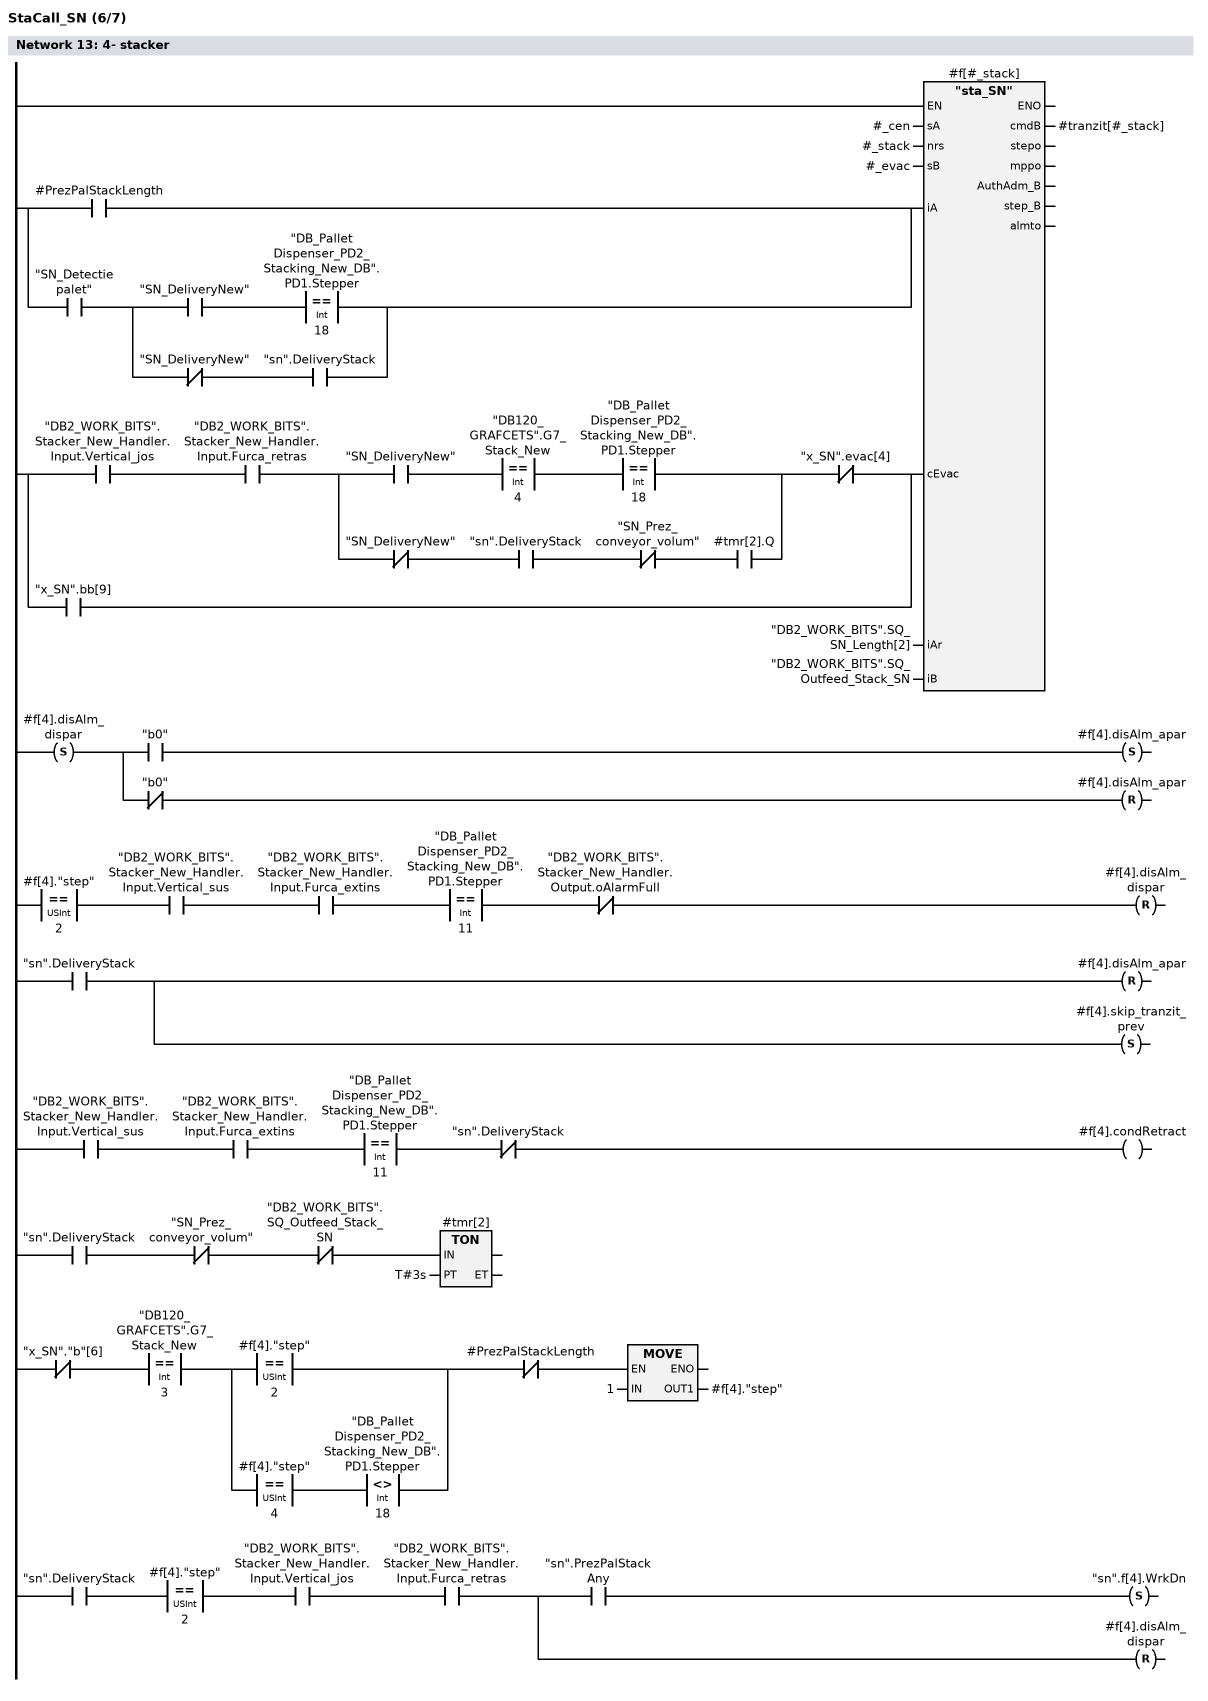
   #f[#_stack](sA := #_cen,   // "sta_SN"
               nrs := #_stack,
               sB := #_evac,
               iA := #PrezPalStackLength OR ("SN_Detectie palet" AND (("SN_DeliveryNew" AND ("DB_PalletDispenser_PD2_Stacking_New_DB".PD1.Stepper = 18)) OR (NOT "SN_DeliveryNew" AND "sn".DeliveryStack))),
               cEvac := ("DB2_WORK_BITS".Stacker_New_Handler.Input.Vertical_jos AND "DB2_WORK_BITS".Stacker_New_Handler.Input.Furca_retras AND (("SN_DeliveryNew" AND ("DB120_GRAFCETS".G7_Stack_New = 4) AND ("DB_PalletDispenser_PD2_Stacking_New_DB".PD1.Stepper = 18)) OR (NOT "SN_DeliveryNew" AND "sn".DeliveryStack AND NOT "SN_Prez_conveyor_volum" AND #tmr[2].Q)) AND NOT "x_SN".evac[4]) OR "x_SN".bb[9],
               iAr := "DB2_WORK_BITS".SQ_SN_Length[2],
               iB := "DB2_WORK_BITS".SQ_Outfeed_Stack_SN,
               cmdB => #tranzit[#_stack]);
   #f[4].disAlm_dispar := TRUE;
   IF "b0" THEN #f[4].disAlm_apar := TRUE; END_IF;
   IF NOT "b0" THEN #f[4].disAlm_apar := FALSE; END_IF;
   IF (#f[4]."step" = 2) AND "DB2_WORK_BITS".Stacker_New_Handler.Input.Vertical_sus AND "DB2_WORK_BITS".Stacker_New_Handler.Input.Furca_extins AND ("DB_PalletDispenser_PD2_Stacking_New_DB".PD1.Stepper = 11) AND NOT "DB2_WORK_BITS".Stacker_New_Handler.Output.oAlarmFull THEN
       #f[4].disAlm_dispar := FALSE;
   END_IF;
   IF "sn".DeliveryStack THEN
       #f[4].disAlm_apar := FALSE;
       #f[4].skip_tranzit_prev := TRUE;
   END_IF;
   #f[4].condRetract := "DB2_WORK_BITS".Stacker_New_Handler.Input.Vertical_sus AND "DB2_WORK_BITS".Stacker_New_Handler.Input.Furca_extins AND ("DB_PalletDispenser_PD2_Stacking_New_DB".PD1.Stepper = 11) AND NOT "sn".DeliveryStack;
   #tmr[2].TON(IN := "sn".DeliveryStack AND NOT "SN_Prez_conveyor_volum" AND NOT "DB2_WORK_BITS".SQ_Outfeed_Stack_SN,
               PT := T#3s);
   IF NOT "x_SN"."b"[6] AND ("DB120_GRAFCETS".G7_Stack_New = 3) AND ((#f[4]."step" = 2) OR ((#f[4]."step" = 4) AND ("DB_PalletDispenser_PD2_Stacking_New_DB".PD1.Stepper <> 18))) AND NOT #PrezPalStackLength THEN
       #f[4]."step" := 1;
   END_IF;
   #_w1 := "sn".DeliveryStack AND (#f[4]."step" = 2) AND "DB2_WORK_BITS".Stacker_New_Handler.Input.Vertical_jos AND "DB2_WORK_BITS".Stacker_New_Handler.Input.Furca_retras;
   IF #_w1 AND "sn".PrezPalStackAny THEN "sn".f[4].WrkDn := TRUE; END_IF;
   IF #_w1 THEN #f[4].disAlm_dispar := FALSE; END_IF;
END_REGION

REGION Network 14: 5- evac
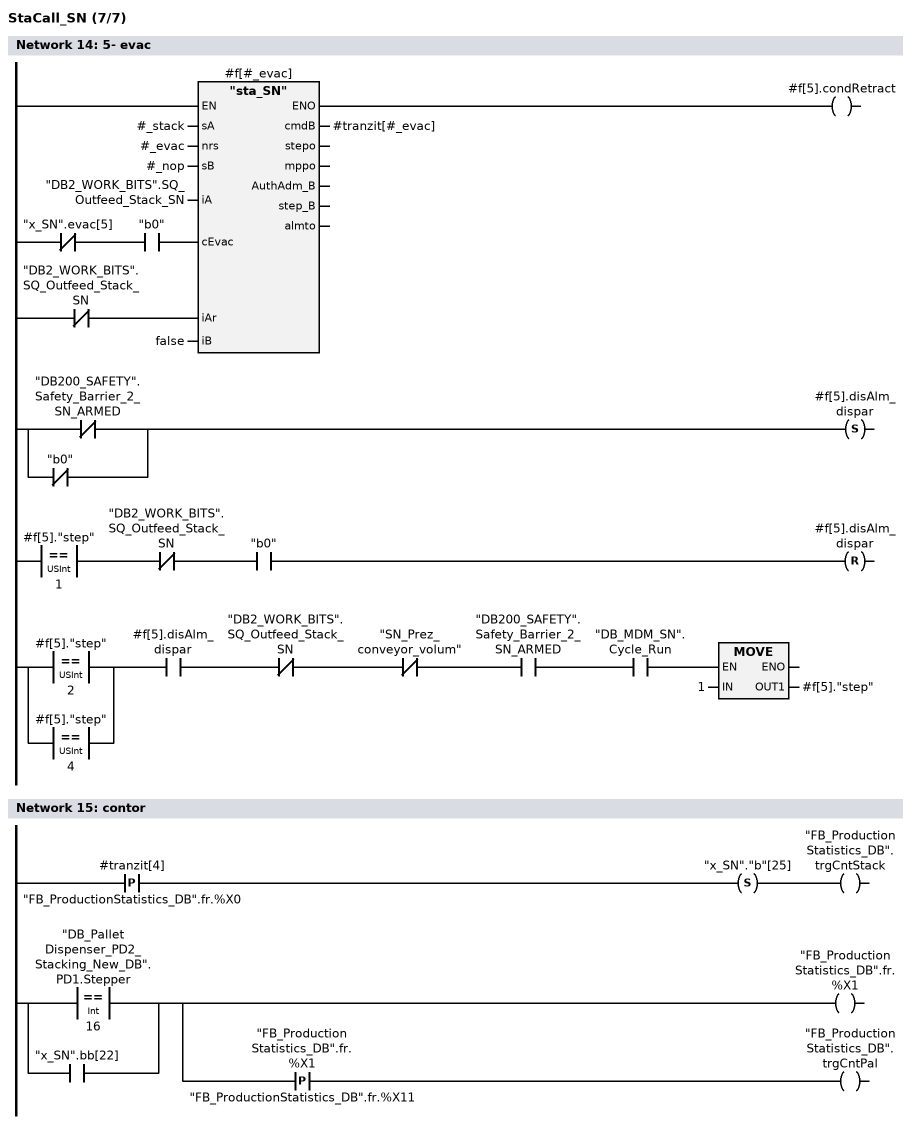
   RUNG wire#powerrail
      #f[#_evac](cEvac := wire#w1, iAr := wire#w2, sA := #_stack, nrs := #_evac, sB := #_nop, iA := "DB2_WORK_BITS".SQ_Outfeed_Stack_SN, iB := false, cmdB => #tranzit[#_evac], stepo =>, mppo =>, AuthAdm_B =>, step_B =>, almto =>)
      Coil( #f[5].condRetract )
   END_RUNG
   RUNG wire#powerrail
      I_Contact( "x_SN".evac[5] )
      Contact( "b0" )
   END_RUNG wire#w1
   RUNG wire#powerrail
      I_Contact( "DB2_WORK_BITS".SQ_Outfeed_Stack_SN )
   END_RUNG wire#w2
   RUNG wire#powerrail
      I_Contact( "DB200_SAFETY".Safety_Barrier_2_SN_ARMED )
      wire#w3
      S_Coil( #f[5].disAlm_dispar )
   END_RUNG
   RUNG wire#powerrail
      I_Contact( "b0" )
   END_RUNG wire#w3
   RUNG wire#powerrail
      { S7_Templates := "SrcType := USInt" } EQ_Contact(in1 := #f[5]."step", in2 := 1)
      I_Contact( "DB2_WORK_BITS".SQ_Outfeed_Stack_SN )
      Contact( "b0" )
      R_Coil( #f[5].disAlm_dispar )
   END_RUNG
   RUNG wire#powerrail
      { S7_Templates := "SrcType := USInt" } EQ_Contact(in1 := #f[5]."step", in2 := 2)
      wire#w4
      Contact( #f[5].disAlm_dispar )
      I_Contact( "DB2_WORK_BITS".SQ_Outfeed_Stack_SN )
      I_Contact( "SN_Prez_conveyor_volum" )
      Contact( "DB200_SAFETY".Safety_Barrier_2_SN_ARMED )
      Contact( "DB_MDM_SN".Cycle_Run )
      Move(in := 1, out1 => #f[5]."step")
   END_RUNG
   RUNG wire#powerrail
      { S7_Templates := "SrcType := USInt" } EQ_Contact(in1 := #f[5]."step", in2 := 4)
   END_RUNG wire#w4
   // the same network as SCL:
   #f[#_evac](sA := #_stack,   // "sta_SN"
              nrs := #_evac,
              sB := #_nop,
              iA := "DB2_WORK_BITS".SQ_Outfeed_Stack_SN,
              cEvac := NOT "x_SN".evac[5] AND "b0",
              iAr := NOT "DB2_WORK_BITS".SQ_Outfeed_Stack_SN,
              iB := false,
              cmdB => #tranzit[#_evac],
              ENO => #_w1);
   #f[5].condRetract := #_w1;
   IF NOT "DB200_SAFETY".Safety_Barrier_2_SN_ARMED OR NOT "b0" THEN #f[5].disAlm_dispar := TRUE; END_IF;
   IF (#f[5]."step" = 1) AND NOT "DB2_WORK_BITS".SQ_Outfeed_Stack_SN AND "b0" THEN
       #f[5].disAlm_dispar := FALSE;
   END_IF;
   IF ((#f[5]."step" = 2) OR (#f[5]."step" = 4)) AND #f[5].disAlm_dispar AND NOT "DB2_WORK_BITS".SQ_Outfeed_Stack_SN AND NOT "SN_Prez_conveyor_volum" AND "DB200_SAFETY".Safety_Barrier_2_SN_ARMED AND "DB_MDM_SN".Cycle_Run THEN
       #f[5]."step" := 1;
   END_IF;
END_REGION

REGION Network 15: contor
   RUNG wire#powerrail
      P_Contact(operand := #tranzit[4], bit := "FB_ProductionStatistics_DB".fr.%X0)
      S_Coil( "x_SN"."b"[25] )
      Coil( "FB_ProductionStatistics_DB".trgCntStack )
   END_RUNG
   RUNG wire#powerrail
      { S7_Templates := "SrcType := Int" } EQ_Contact(in1 := "DB_PalletDispenser_PD2_Stacking_New_DB".PD1.Stepper, in2 := 16)
      wire#w1
      Coil( "FB_ProductionStatistics_DB".fr.%X1 )
   END_RUNG
   RUNG wire#powerrail
      Contact( "x_SN".bb[22] )
   END_RUNG wire#w1
   RUNG wire#w1
      P_Contact(operand := "FB_ProductionStatistics_DB".fr.%X1, bit := "FB_ProductionStatistics_DB".fr.%X11)
      Coil( "FB_ProductionStatistics_DB".trgCntPal )
   END_RUNG
   // the same network as SCL:
   #_w1 := #tranzit[4] AND NOT "FB_ProductionStatistics_DB".fr.%X0;   // rising edge of #tranzit[4]
   "FB_ProductionStatistics_DB".fr.%X0 := #tranzit[4];
   IF #_w1 THEN "x_SN"."b"[25] := TRUE; END_IF;
   "FB_ProductionStatistics_DB".trgCntStack := #_w1;
   "FB_ProductionStatistics_DB".fr.%X1 := ("DB_PalletDispenser_PD2_Stacking_New_DB".PD1.Stepper = 16) OR "x_SN".bb[22];
   #_w2 := "FB_ProductionStatistics_DB".fr.%X1 AND "FB_ProductionStatistics_DB".fr.%X1 AND NOT "FB_ProductionStatistics_DB".fr.%X11;   // rising edge of "FB_ProductionStatistics_DB".fr.%X1
   "FB_ProductionStatistics_DB".fr.%X11 := "FB_ProductionStatistics_DB".fr.%X1;
   "FB_ProductionStatistics_DB".trgCntPal := #_w2;
END_REGION
END_FUNCTION_BLOCK

FUNCTION_BLOCK "sta_SN"   // FB16, LAD
{ S7_Optimized_Access := 'TRUE' }
VERSION : 0.1
   VAR_INPUT
      sA : USInt;   // statie Admit
      nrs : USInt;   // statie crt
      sB : USInt;   // statie Evac
      iA : Bool;   // conditie Admit
      cEvac : Bool;
      iAr : Bool;   // cond Release
      iB : Bool;   // cond Evac
   END_VAR
   VAR_OUTPUT
      cmdB : Bool;
      stepo : USInt;
      mppo : Bool;
      AuthAdm_B : Bool;
      step_B : USInt;
      almto : USInt;
   END_VAR
   VAR
      "step" : USInt;
      stepv : USInt;
      mpp : Bool;
      alm_apar : Bool;
      alm_disapear : Bool;
      alm_tmt : Bool;
      alm_release : Bool;
      AuthAdmit : Bool;
      AuthEvacEx : Bool;
      almt : Bool;
      WrkDn : Bool;
      condRetract : Bool;
      skip_tranzit_prev : Bool;
      product_disapear_confirmed : Bool;
      transit_end_confirmed : Bool;
      tim_alm : Array[1..6] of IEC_TIMER;
      HMI_stat_s : USInt;
      disAlm_Tmt : Bool;
      disAlm_dispar : Bool;
      disAlm_apar : Bool;
      disAlmRls : Bool;
      HMI_stat_t : USInt;
      tranzit_mem : Bool;
      cycle : Bool;
      almw : Word;
      HMI_statT : USInt;
      HMI_statS : USInt;
      tr : USInt;
      AlarmW : Word;
   END_VAR
   VAR_TEMP
      tmpui : SInt;
   END_VAR
   VAR CONSTANT
      b0 : Bool;
   END_VAR
   VAR_TEMP   // added for the SCL form of the ladder/FBD networks
      _w1 : Bool;
      _w2 : Bool;
      _w3 : Bool;
   END_VAR
BEGIN

REGION Network 1: first cycle
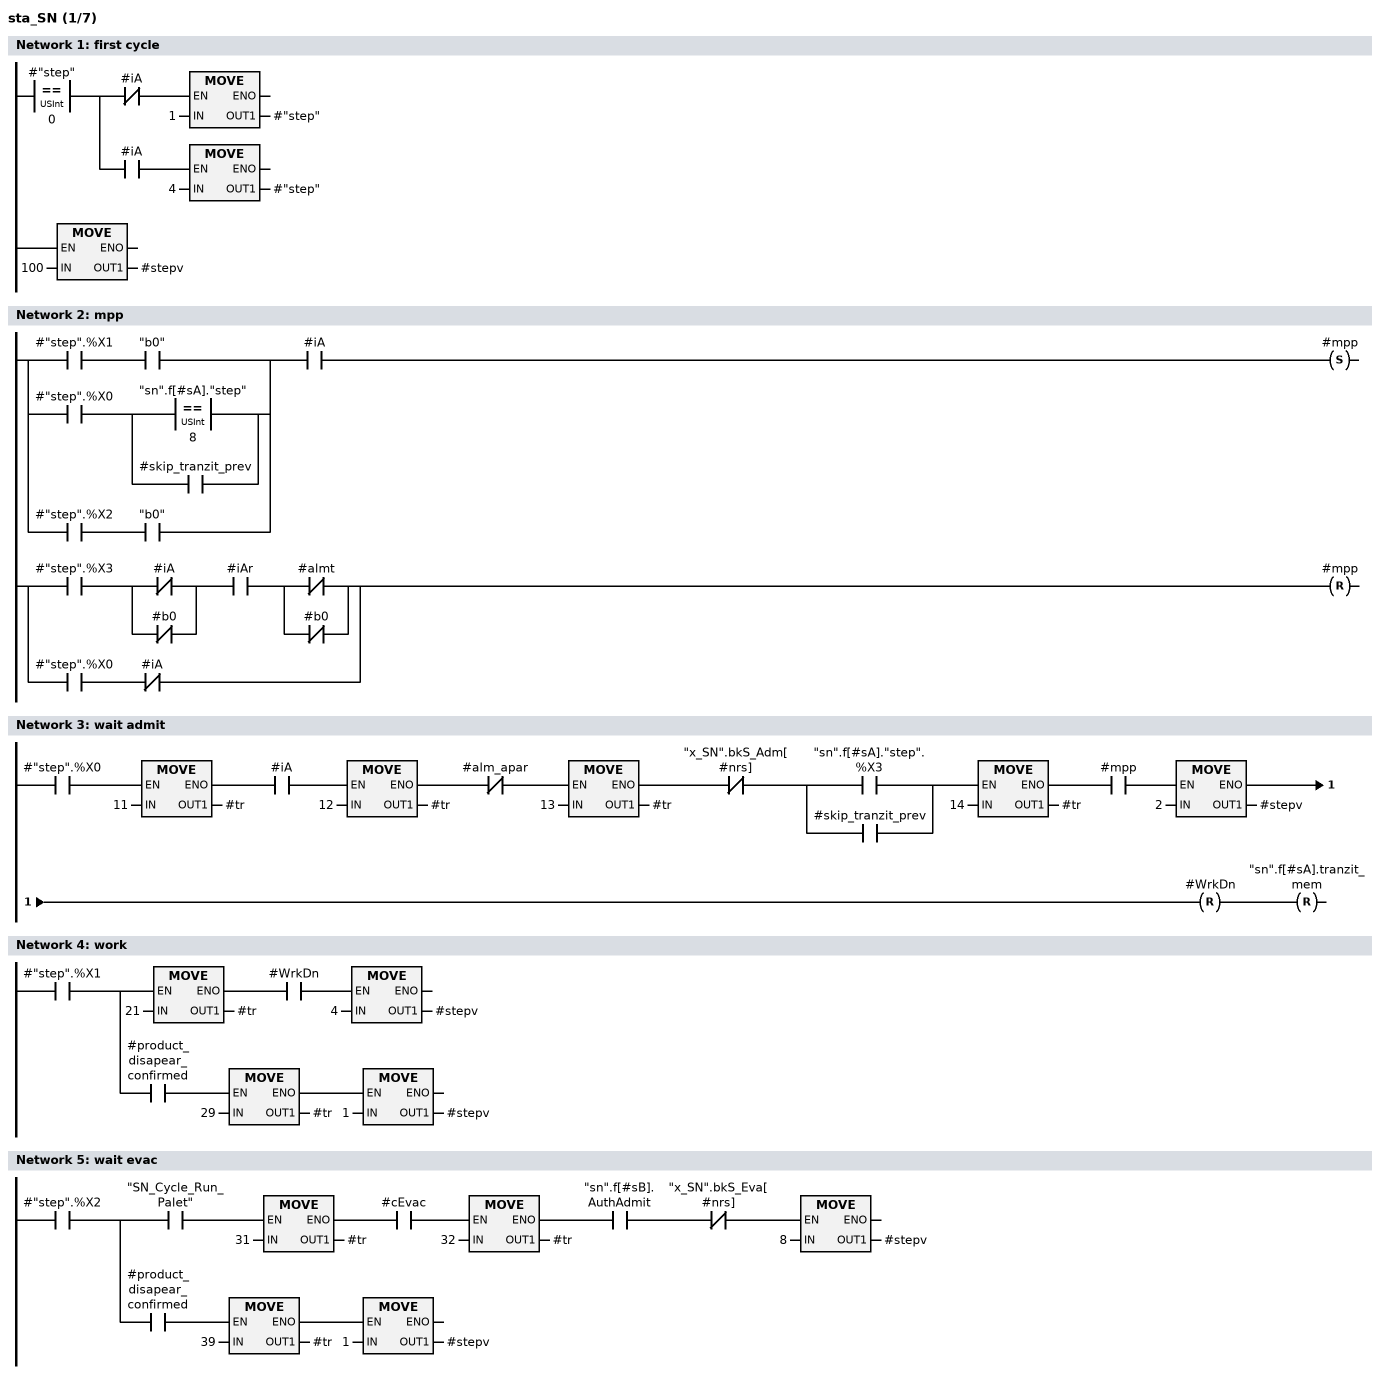
   RUNG wire#powerrail
      { S7_Templates := "SrcType := USInt" } EQ_Contact(in1 := #"step", in2 := 0)
      wire#w1
      I_Contact( #iA )
      Move(in := 1, out1 => #"step")
   END_RUNG
   RUNG wire#w1
      Contact( #iA )
      Move(in := 4, out1 => #"step")
   END_RUNG
   RUNG wire#powerrail
      Move(in := 100, out1 => #stepv)
   END_RUNG
   // the same network as SCL:
   #_w1 := #"step" = 0;
   IF #_w1 AND NOT #iA THEN #"step" := 1; END_IF;
   IF #_w1 AND #iA THEN #"step" := 4; END_IF;
   #stepv := 100;
END_REGION

REGION Network 2: mpp
   RUNG wire#powerrail
      Contact( #"step".%X1 )
      Contact( "b0" )
      wire#w1
      Contact( #iA )
      S_Coil( #mpp )
   END_RUNG
   RUNG wire#powerrail
      Contact( #"step".%X0 )
      wire#w2
      { S7_Templates := "SrcType := USInt" } EQ_Contact(in1 := "sn".f[#sA]."step", in2 := 8)
   END_RUNG wire#w1
   RUNG wire#w2
      Contact( #skip_tranzit_prev )
   END_RUNG wire#w1
   RUNG wire#powerrail
      Contact( #"step".%X2 )
      Contact( "b0" )
   END_RUNG wire#w1
   RUNG wire#powerrail
      Contact( #"step".%X3 )
      wire#w3
      I_Contact( #iA )
      wire#w4
      Contact( #iAr )
      wire#w5
      I_Contact( #almt )
      wire#w6
      R_Coil( #mpp )
   END_RUNG
   RUNG wire#w3
      I_Contact( #b0 )
   END_RUNG wire#w4
   RUNG wire#w5
      I_Contact( #b0 )
   END_RUNG wire#w6
   RUNG wire#powerrail
      Contact( #"step".%X0 )
      I_Contact( #iA )
   END_RUNG wire#w6
   // the same network as SCL:
   IF ((#"step".%X1 AND "b0") OR (#"step".%X0 AND (("sn".f[#sA]."step" = 8) OR #skip_tranzit_prev)) OR (#"step".%X2 AND "b0")) AND #iA THEN
       #mpp := TRUE;
   END_IF;
   IF (#"step".%X3 AND (NOT #iA OR NOT #b0) AND #iAr AND (NOT #almt OR NOT #b0)) OR (#"step".%X0 AND NOT #iA) THEN
       #mpp := FALSE;
   END_IF;
END_REGION

REGION Network 3: wait admit
   RUNG wire#powerrail
      Contact( #"step".%X0 )
      Move(in := 11, out1 => #tr)
      Contact( #iA )
      Move(in := 12, out1 => #tr)
      I_Contact( #alm_apar )
      Move(in := 13, out1 => #tr)
      I_Contact( "x_SN".bkS_Adm[#nrs] )
      wire#w1
      Contact( "sn".f[#sA]."step".%X3 )
      wire#w2
      Move(in := 14, out1 => #tr)
      Contact( #mpp )
      Move(in := 2, out1 => #stepv)
      R_Coil( #WrkDn )
      R_Coil( "sn".f[#sA].tranzit_mem )
   END_RUNG
   RUNG wire#w1
      Contact( #skip_tranzit_prev )
   END_RUNG wire#w2
   // the same network as SCL:
   IF #"step".%X0 THEN #tr := 11; END_IF;
   #_w1 := #"step".%X0 AND #iA;
   IF #_w1 THEN #tr := 12; END_IF;
   #_w2 := #_w1 AND NOT #alm_apar;
   IF #_w2 THEN #tr := 13; END_IF;
   #_w3 := #_w2 AND NOT "x_SN".bkS_Adm[#nrs] AND ("sn".f[#sA]."step".%X3 OR #skip_tranzit_prev);
   IF #_w3 THEN #tr := 14; END_IF;
   IF #_w3 AND #mpp THEN
       #stepv := 2;
       #WrkDn := FALSE;
       "sn".f[#sA].tranzit_mem := FALSE;
   END_IF;
END_REGION

REGION Network 4: work
   RUNG wire#powerrail
      Contact( #"step".%X1 )
      wire#w1
      Move(in := 21, out1 => #tr)
      Contact( #WrkDn )
      Move(in := 4, out1 => #stepv)
   END_RUNG
   RUNG wire#w1
      Contact( #product_disapear_confirmed )
      Move(in := 29, out1 => #tr)
      Move(in := 1, out1 => #stepv)
   END_RUNG
   // the same network as SCL:
   IF #"step".%X1 THEN #tr := 21; END_IF;
   IF #"step".%X1 AND #WrkDn THEN #stepv := 4; END_IF;
   IF #"step".%X1 AND #product_disapear_confirmed THEN
       #tr := 29;
       #stepv := 1;
   END_IF;
END_REGION

REGION Network 5: wait evac
   RUNG wire#powerrail
      Contact( #"step".%X2 )
      wire#w1
      Contact( "SN_Cycle_Run_Palet" )
      Move(in := 31, out1 => #tr)
      Contact( #cEvac )
      Move(in := 32, out1 => #tr)
      Contact( "sn".f[#sB].AuthAdmit )
      I_Contact( "x_SN".bkS_Eva[#nrs] )
      Move(in := 8, out1 => #stepv)
   END_RUNG
   RUNG wire#w1
      Contact( #product_disapear_confirmed )
      Move(in := 39, out1 => #tr)
      Move(in := 1, out1 => #stepv)
   END_RUNG
   // the same network as SCL:
   #_w1 := #"step".%X2 AND "SN_Cycle_Run_Palet";
   IF #_w1 THEN #tr := 31; END_IF;
   #_w2 := #_w1 AND #cEvac;
   IF #_w2 THEN #tr := 32; END_IF;
   IF #_w2 AND "sn".f[#sB].AuthAdmit AND NOT "x_SN".bkS_Eva[#nrs] THEN #stepv := 8; END_IF;
   IF #"step".%X2 AND #product_disapear_confirmed THEN
       #tr := 39;
       #stepv := 1;
   END_IF;
END_REGION

REGION Network 6: evac
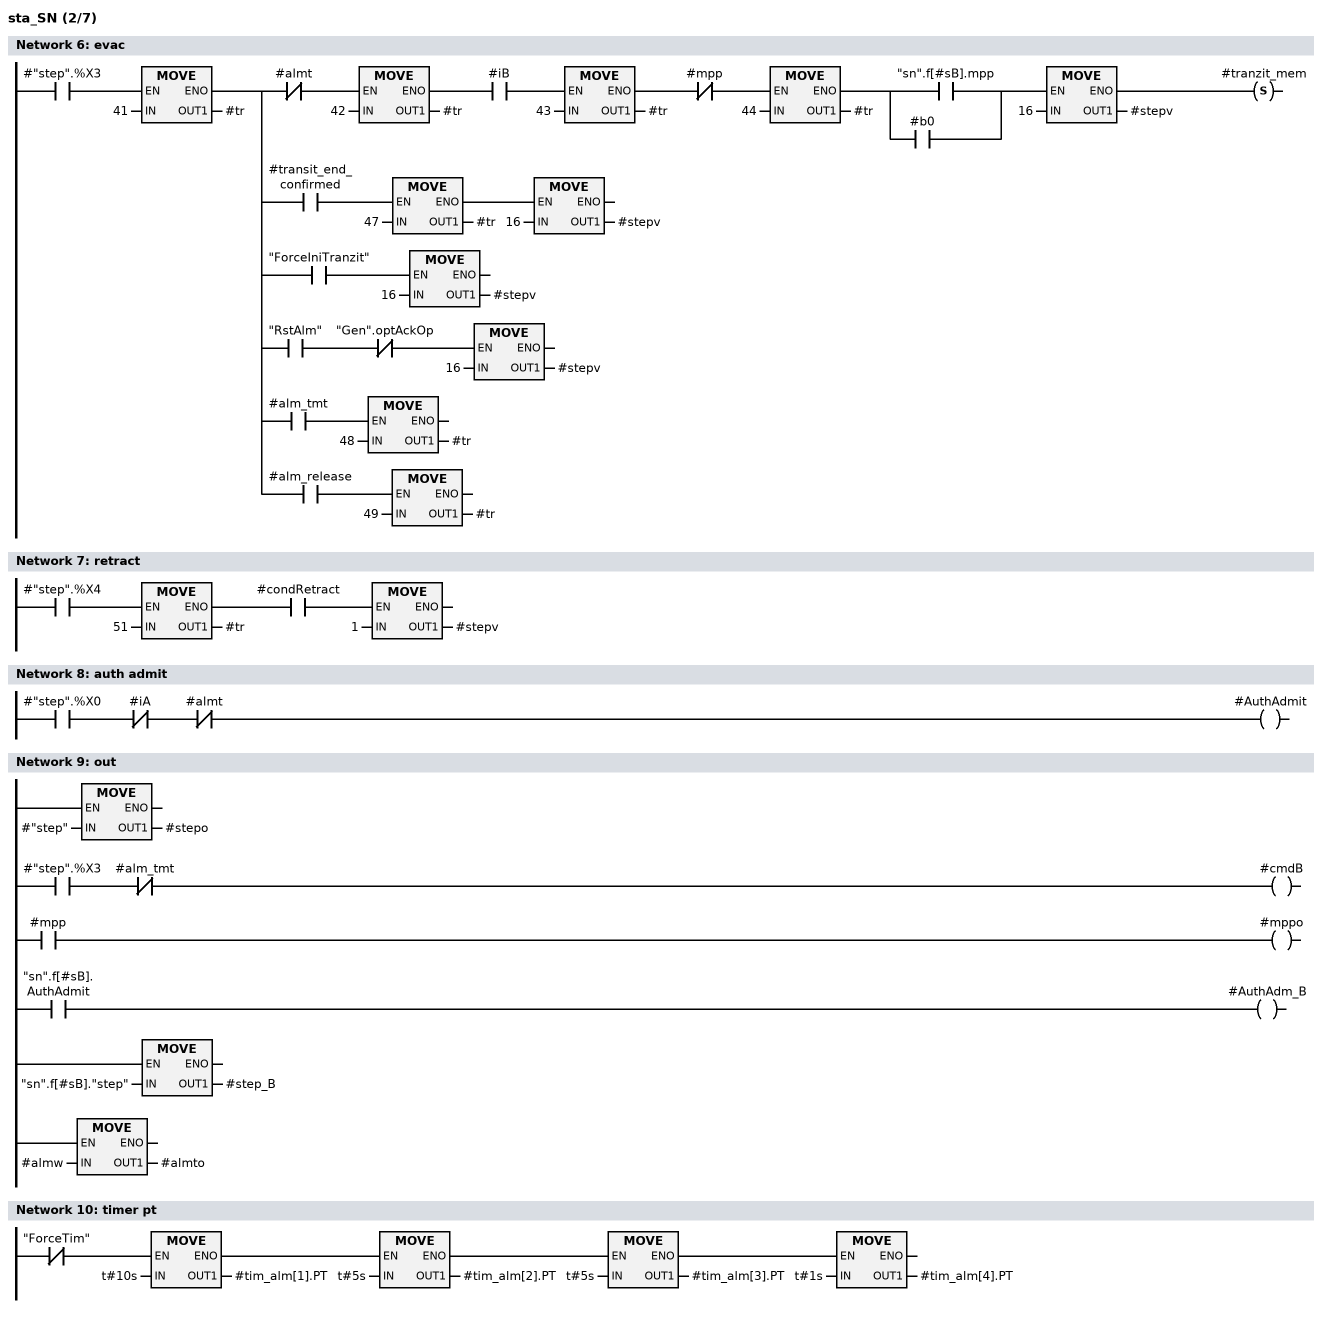
   RUNG wire#powerrail
      Contact( #"step".%X3 )
      Move(in := 41, out1 => #tr)
      wire#w1
      I_Contact( #almt )
      Move(in := 42, out1 => #tr)
      Contact( #iB )
      Move(in := 43, out1 => #tr)
      I_Contact( #mpp )
      Move(in := 44, out1 => #tr)
      wire#w2
      Contact( "sn".f[#sB].mpp )
      wire#w3
      Move(in := 16, out1 => #stepv)
      S_Coil( #tranzit_mem )
   END_RUNG
   RUNG wire#w2
      Contact( #b0 )
   END_RUNG wire#w3
   RUNG wire#w1
      Contact( #transit_end_confirmed )
      Move(in := 47, out1 => #tr)
      Move(in := 16, out1 => #stepv)
   END_RUNG
   RUNG wire#w1
      Contact( "ForceIniTranzit" )
      Move(in := 16, out1 => #stepv)
   END_RUNG
   RUNG wire#w1
      Contact( "RstAlm" )
      I_Contact( "Gen".optAckOp )
      Move(in := 16, out1 => #stepv)
   END_RUNG
   RUNG wire#w1
      Contact( #alm_tmt )
      Move(in := 48, out1 => #tr)
   END_RUNG
   RUNG wire#w1
      Contact( #alm_release )
      Move(in := 49, out1 => #tr)
   END_RUNG
   // the same network as SCL:
   IF #"step".%X3 THEN #tr := 41; END_IF;
   #_w1 := #"step".%X3 AND NOT #almt;
   IF #_w1 THEN #tr := 42; END_IF;
   #_w2 := #_w1 AND #iB;
   IF #_w2 THEN #tr := 43; END_IF;
   #_w3 := #_w2 AND NOT #mpp;
   IF #_w3 THEN #tr := 44; END_IF;
   IF #_w3 AND ("sn".f[#sB].mpp OR #b0) THEN
       #stepv := 16;
       #tranzit_mem := TRUE;
   END_IF;
   IF #"step".%X3 AND #transit_end_confirmed THEN
       #tr := 47;
       #stepv := 16;
   END_IF;
   IF #"step".%X3 AND "ForceIniTranzit" THEN #stepv := 16; END_IF;
   IF #"step".%X3 AND "RstAlm" AND NOT "Gen".optAckOp THEN #stepv := 16; END_IF;
   IF #"step".%X3 AND #alm_tmt THEN #tr := 48; END_IF;
   IF #"step".%X3 AND #alm_release THEN #tr := 49; END_IF;
END_REGION

REGION Network 7: retract
   RUNG wire#powerrail
      Contact( #"step".%X4 )
      Move(in := 51, out1 => #tr)
      Contact( #condRetract )
      Move(in := 1, out1 => #stepv)
   END_RUNG
   // the same network as SCL:
   IF #"step".%X4 THEN #tr := 51; END_IF;
   IF #"step".%X4 AND #condRetract THEN #stepv := 1; END_IF;
END_REGION

REGION Network 8: auth admit
   RUNG wire#powerrail
      Contact( #"step".%X0 )
      I_Contact( #iA )
      I_Contact( #almt )
      Coil( #AuthAdmit )
   END_RUNG
   // the same network as SCL:
   #AuthAdmit := #"step".%X0 AND NOT #iA AND NOT #almt;
END_REGION

REGION Network 9: out
   RUNG wire#powerrail
      Move(in := #"step", out1 => #stepo)
   END_RUNG
   RUNG wire#powerrail
      Contact( #"step".%X3 )
      I_Contact( #alm_tmt )
      Coil( #cmdB )
   END_RUNG
   RUNG wire#powerrail
      Contact( #mpp )
      Coil( #mppo )
   END_RUNG
   RUNG wire#powerrail
      Contact( "sn".f[#sB].AuthAdmit )
      Coil( #AuthAdm_B )
   END_RUNG
   RUNG wire#powerrail
      Move(in := "sn".f[#sB]."step", out1 => #step_B)
   END_RUNG
   RUNG wire#powerrail
      Move(in := #almw, out1 => #almto)
   END_RUNG
   // the same network as SCL:
   #stepo := #"step";
   #cmdB := #"step".%X3 AND NOT #alm_tmt;
   #mppo := #mpp;
   #AuthAdm_B := "sn".f[#sB].AuthAdmit;
   #step_B := "sn".f[#sB]."step";
   #almto := #almw;
END_REGION

REGION Network 10: timer pt
   RUNG wire#powerrail
      I_Contact( "ForceTim" )
      Move(in := t#10s, out1 => #tim_alm[1].PT)
      Move(in := t#5s, out1 => #tim_alm[2].PT)
      Move(in := t#5s, out1 => #tim_alm[3].PT)
      Move(in := t#1s, out1 => #tim_alm[4].PT)
   END_RUNG
   // the same network as SCL:
   IF NOT "ForceTim" THEN
       #tim_alm[1].PT := t#10s;
       #tim_alm[2].PT := t#5s;
       #tim_alm[3].PT := t#5s;
       #tim_alm[4].PT := t#1s;
   END_IF;
END_REGION

REGION Network 11: rst all
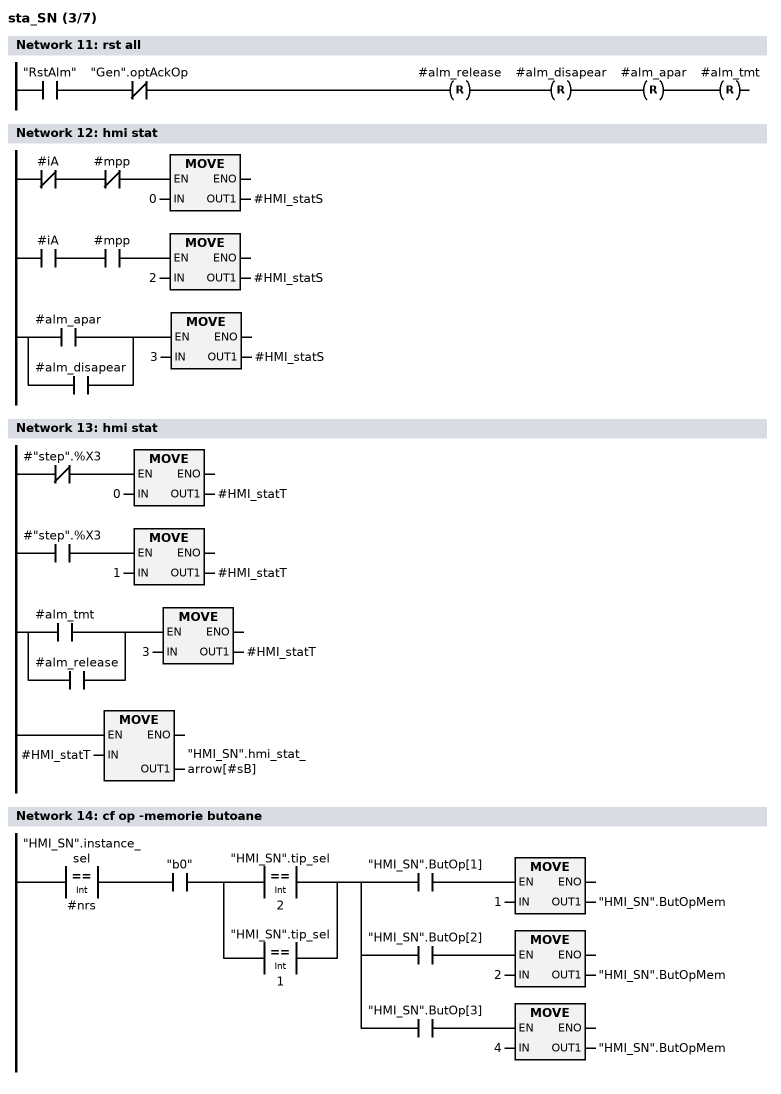
   RUNG wire#powerrail
      Contact( "RstAlm" )
      I_Contact( "Gen".optAckOp )
      R_Coil( #alm_release )
      R_Coil( #alm_disapear )
      R_Coil( #alm_apar )
      R_Coil( #alm_tmt )
   END_RUNG
   // the same network as SCL:
   IF "RstAlm" AND NOT "Gen".optAckOp THEN
       #alm_release := FALSE;
       #alm_disapear := FALSE;
       #alm_apar := FALSE;
       #alm_tmt := FALSE;
   END_IF;
END_REGION

REGION Network 12: hmi stat
   RUNG wire#powerrail
      I_Contact( #iA )
      I_Contact( #mpp )
      Move(in := 0, out1 => #HMI_statS)
   END_RUNG
   RUNG wire#powerrail
      Contact( #iA )
      Contact( #mpp )
      Move(in := 2, out1 => #HMI_statS)
   END_RUNG
   RUNG wire#powerrail
      Contact( #alm_apar )
      wire#w1
      Move(in := 3, out1 => #HMI_statS)
   END_RUNG
   RUNG wire#powerrail
      Contact( #alm_disapear )
   END_RUNG wire#w1
   // the same network as SCL:
   IF NOT #iA AND NOT #mpp THEN #HMI_statS := 0; END_IF;
   IF #iA AND #mpp THEN #HMI_statS := 2; END_IF;
   IF #alm_apar OR #alm_disapear THEN #HMI_statS := 3; END_IF;
END_REGION

REGION Network 13: hmi stat
   RUNG wire#powerrail
      I_Contact( #"step".%X3 )
      Move(in := 0, out1 => #HMI_statT)
   END_RUNG
   RUNG wire#powerrail
      Contact( #"step".%X3 )
      Move(in := 1, out1 => #HMI_statT)
   END_RUNG
   RUNG wire#powerrail
      Contact( #alm_tmt )
      wire#w1
      Move(in := 3, out1 => #HMI_statT)
   END_RUNG
   RUNG wire#powerrail
      Contact( #alm_release )
   END_RUNG wire#w1
   RUNG wire#powerrail
      Move(in := #HMI_statT, out1 => "HMI_SN".hmi_stat_arrow[#sB])
   END_RUNG
   // the same network as SCL:
   IF NOT #"step".%X3 THEN #HMI_statT := 0; END_IF;
   IF #"step".%X3 THEN #HMI_statT := 1; END_IF;
   IF #alm_tmt OR #alm_release THEN #HMI_statT := 3; END_IF;
   "HMI_SN".hmi_stat_arrow[#sB] := #HMI_statT;
END_REGION

REGION Network 14: cf op -memorie butoane
   RUNG wire#powerrail
      { S7_Templates := "SrcType := Int" } EQ_Contact(in1 := "HMI_SN".instance_sel, in2 := #nrs)
      Contact( "b0" )
      wire#w1
      { S7_Templates := "SrcType := Int" } EQ_Contact(in1 := "HMI_SN".tip_sel, in2 := 2)
      wire#w2
      Contact( "HMI_SN".ButOp[1] )
      Move(in := 1, out1 => "HMI_SN".ButOpMem)
   END_RUNG
   RUNG wire#w1
      { S7_Templates := "SrcType := Int" } EQ_Contact(in1 := "HMI_SN".tip_sel, in2 := 1)
   END_RUNG wire#w2
   RUNG wire#w2
      Contact( "HMI_SN".ButOp[2] )
      Move(in := 2, out1 => "HMI_SN".ButOpMem)
   END_RUNG
   RUNG wire#w2
      Contact( "HMI_SN".ButOp[3] )
      Move(in := 4, out1 => "HMI_SN".ButOpMem)
   END_RUNG
   // the same network as SCL:
   #_w1 := ("HMI_SN".instance_sel = #nrs) AND "b0" AND (("HMI_SN".tip_sel = 2) OR ("HMI_SN".tip_sel = 1));
   IF #_w1 AND "HMI_SN".ButOp[1] THEN "HMI_SN".ButOpMem := 1; END_IF;
   IF #_w1 AND "HMI_SN".ButOp[2] THEN "HMI_SN".ButOpMem := 2; END_IF;
   IF #_w1 AND "HMI_SN".ButOp[3] THEN "HMI_SN".ButOpMem := 4; END_IF;
END_REGION

REGION Network 15: cf op alm tmt / release
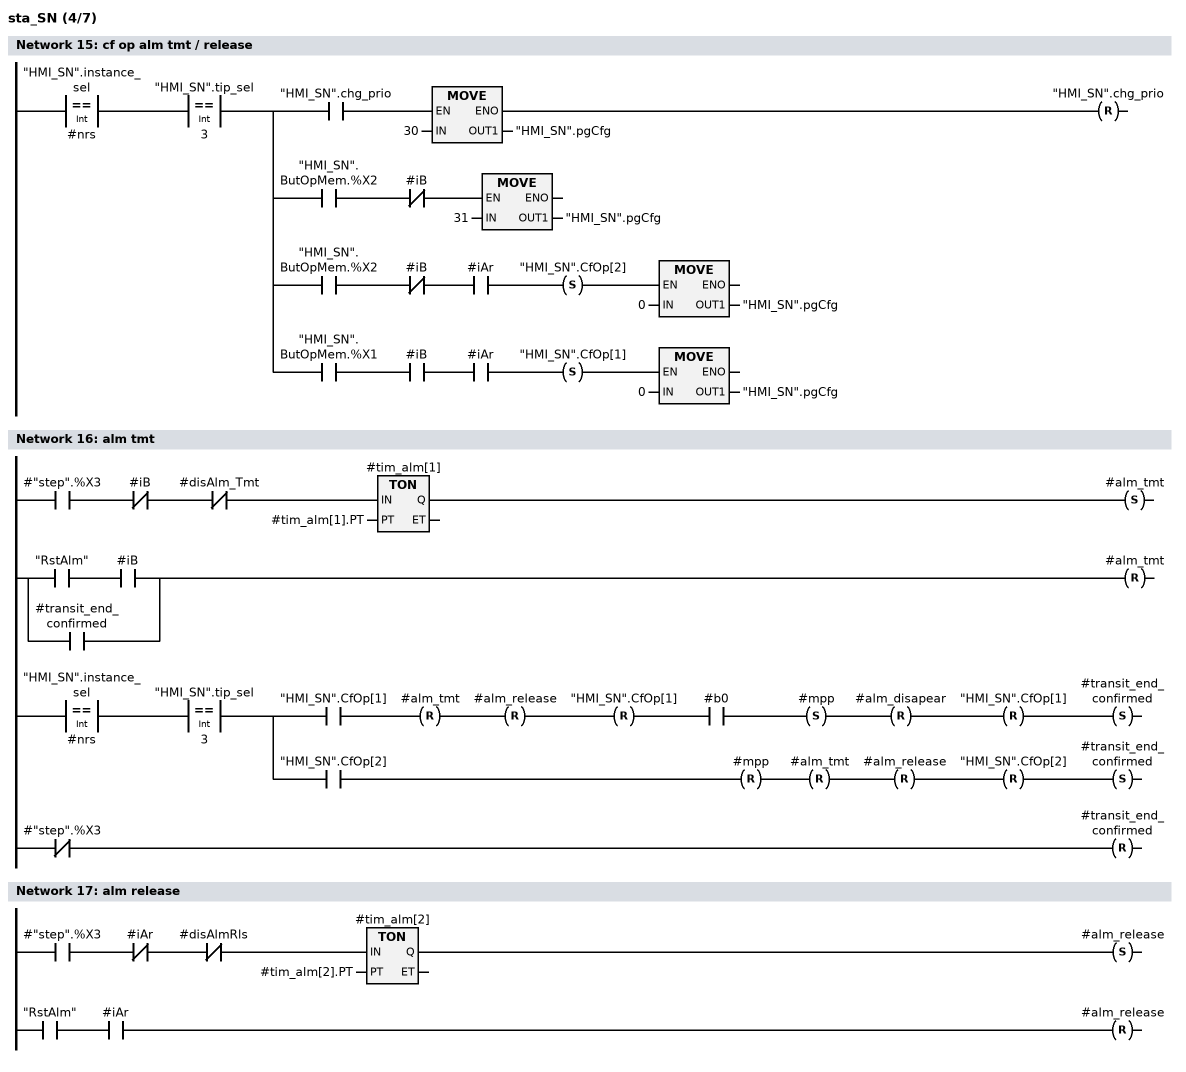
   RUNG wire#powerrail
      { S7_Templates := "SrcType := Int" } EQ_Contact(in1 := "HMI_SN".instance_sel, in2 := #nrs)
      { S7_Templates := "SrcType := Int" } EQ_Contact(in1 := "HMI_SN".tip_sel, in2 := 3)
      wire#w1
      Contact( "HMI_SN".chg_prio )
      Move(in := 30, out1 => "HMI_SN".pgCfg)
      R_Coil( "HMI_SN".chg_prio )
   END_RUNG
   RUNG wire#w1
      Contact( "HMI_SN".ButOpMem.%X2 )
      I_Contact( #iB )
      Move(in := 31, out1 => "HMI_SN".pgCfg)
   END_RUNG
   RUNG wire#w1
      Contact( "HMI_SN".ButOpMem.%X2 )
      I_Contact( #iB )
      Contact( #iAr )
      S_Coil( "HMI_SN".CfOp[2] )
      Move(in := 0, out1 => "HMI_SN".pgCfg)
   END_RUNG
   RUNG wire#w1
      Contact( "HMI_SN".ButOpMem.%X1 )
      Contact( #iB )
      Contact( #iAr )
      S_Coil( "HMI_SN".CfOp[1] )
      Move(in := 0, out1 => "HMI_SN".pgCfg)
   END_RUNG
   // the same network as SCL:
   #_w1 := ("HMI_SN".instance_sel = #nrs) AND ("HMI_SN".tip_sel = 3);
   IF #_w1 AND "HMI_SN".chg_prio THEN
       "HMI_SN".pgCfg := 30;
       "HMI_SN".chg_prio := FALSE;
   END_IF;
   IF #_w1 AND "HMI_SN".ButOpMem.%X2 AND NOT #iB THEN "HMI_SN".pgCfg := 31; END_IF;
   IF #_w1 AND "HMI_SN".ButOpMem.%X2 AND NOT #iB AND #iAr THEN
       "HMI_SN".CfOp[2] := TRUE;
       "HMI_SN".pgCfg := 0;
   END_IF;
   IF #_w1 AND "HMI_SN".ButOpMem.%X1 AND #iB AND #iAr THEN
       "HMI_SN".CfOp[1] := TRUE;